   "Carrier_65_Status.3" AT %I3600.3 : Bool;   // POSITIONING_COMPLETE
   "Carrier_65_Status.4" AT %I3600.4 : Bool;   // PRODUCTION HOLD
   "Carrier_65_Status.5" AT %I3600.5 : Bool;   // CARRIER MOVING FORWARD
   "Carrier_65_Status.6" AT %I3600.6 : Bool;   // CARRIER MOVING REVERSE
   "Carrier_65_Status.7" AT %I3600.7 : Bool;   // CARRIER FAULT
   "Carrier_65_Status.8" AT %I3601.0 : Bool;   // CRASH DETECT TRIPPED
   "Carrier_65_Status.9" AT %I3601.1 : Bool;
   "Carrier_65_Status.10" AT %I3601.2 : Bool;
   "Carrier_65_Status.11" AT %I3601.3 : Bool;
   "Carrier_65_Status.12" AT %I3601.4 : Bool;
   "Carrier_65_Status.13" AT %I3601.5 : Bool;
   "Carrier_65_Status.14" AT %I3601.6 : Bool;
   "Carrier_65_Status.15" AT %I3601.7 : Bool;
   "Carrier_65_SDCFaultCode" AT %IW3602 : Word;   // SDC FAULT CODE
   "Carrier_65_CarrierPosition" AT %ID3604 : DWord;   // CARRIER POSITION
   "Carrier_65_CarrierNumber" AT %IW3608 : Word;   // CARRIER NUMBER
   "Carrier_65_G120DControlWord" AT %IW3610 : Word;   // G120D_STW1_CONTROL
   "Carrier_65_G120DControlWord.0" AT %I3610.0 : Bool;   // Bit_00_ON
   "Carrier_65_G120DControlWord.1" AT %I3610.1 : Bool;   // Bit_01_AUS2_INH
   "Carrier_65_G120DControlWord.2" AT %I3610.2 : Bool;   // Bit_02_AUS3_STOP
   "Carrier_65_G120DControlWord.3" AT %I3610.3 : Bool;   // Bit_03_EN
   "Carrier_65_G120DControlWord.4" AT %I3610.4 : Bool;   // Bit_04_EN_RAMP
   "Carrier_65_G120DControlWord.5" AT %I3610.5 : Bool;   // Bit_05_START_RAMP
   "Carrier_65_G120DControlWord.6" AT %I3610.6 : Bool;   // Bit_06_SETPOINT
   "Carrier_65_G120DControlWord.7" AT %I3610.7 : Bool;   // Bit_07_RESET
   "Carrier_65_G120DControlWord.8" AT %I3611.0 : Bool;   // Bit_08_JOG_R
   "Carrier_65_G120DControlWord.9" AT %I3611.1 : Bool;   // Bit_09_JOG_L
   "Carrier_65_G120DControlWord.10" AT %I3611.2 : Bool;   // Bit_10_CONTR_PLC
   "Carrier_65_G120DControlWord.11" AT %I3611.3 : Bool;   // Bit_11_REVERSE
   "Carrier_65_G120DControlWord.12" AT %I3611.4 : Bool;   // Bit_12_BRAKE_RELEASE
   "Carrier_65_G120DControlWord.13" AT %I3611.5 : Bool;   // Bit_13_DDS
   "Carrier_65_G120DControlWord.14" AT %I3611.6 : Bool;   // Bit_14_DO0
   "Carrier_65_G120DControlWord.15" AT %I3611.7 : Bool;   // Bit_15_DO1
   "Carrier_65_G120DStatusWord" AT %IW3612 : Word;   // G120D_ZSW1_STATUS
   "Carrier_65_G120DStatusWord.0" AT %I3612.0 : Bool;   // Bit_00_READY_RUN
   "Carrier_65_G120DStatusWord.1" AT %I3612.1 : Bool;   // Bit_01_READY_ON
   "Carrier_65_G120DStatusWord.2" AT %I3612.2 : Bool;   // Bit_02_ENABLE
   "Carrier_65_G120DStatusWord.3" AT %I3612.3 : Bool;   // Bit_03_FAULT
   "Carrier_65_G120DStatusWord.4" AT %I3612.4 : Bool;   // Bit_04_OFF2
   "Carrier_65_G120DStatusWord.5" AT %I3612.5 : Bool;   // Bit_05_OFF3
   "Carrier_65_G120DStatusWord.6" AT %I3612.6 : Bool;   // Bit_06_LOCK_OUT
   "Carrier_65_G120DStatusWord.7" AT %I3612.7 : Bool;   // Bit_07_WARN
   "Carrier_65_G120DStatusWord.8" AT %I3613.0 : Bool;   // Bit_08_NO_DEVIATION
   "Carrier_65_G120DStatusWord.9" AT %I3613.1 : Bool;   // Bit_09_CONTR_PLC
   "Carrier_65_G120DStatusWord.10" AT %I3613.2 : Bool;   // Bit_10_F_MAX
   "Carrier_65_G120DStatusWord.11" AT %I3613.3 : Bool;   // Bit_11_LIMIT_REACHED
   "Carrier_65_G120DStatusWord.12" AT %I3613.4 : Bool;   // Bit_12_BRAKE_OPEN
   "Carrier_65_G120DStatusWord.13" AT %I3613.5 : Bool;   // Bit_13_NO_OVERTEMP
   "Carrier_65_G120DStatusWord.14" AT %I3613.6 : Bool;   // Bit_14_CW_CCW
   "Carrier_65_G120DStatusWord.15" AT %I3613.7 : Bool;   // Bit_15_OVERL
   "Carrier_65_Slot2_Input" AT %IW3614 : Word;   // SLOT 2 INPUT WORD
   "Carrier_65_CrashDetectSW" AT %I3614.0 : Bool;   // CRASH DETECT SW
   "Carrier_65_SpareSafetyInput(2_1)" AT %I3614.1 : Bool;   // SPARE SAFETY INPUT
   "Carrier_65_SpareSafetyInput(2_2)" AT %I3614.2 : Bool;   // SPARE SAFETY INPUT
   "Carrier_65_SpareSafetyInput(2_3)" AT %I3614.3 : Bool;   // SPARE SAFETY INPUT
   "Carrier_65_SpareSafetyInput(2_4)" AT %I3614.4 : Bool;   // SPARE SAFETY INPUT
   "Carrier_65_SpareSafetyInput(2_5)" AT %I3614.5 : Bool;   // SPARE SAFETY INPUT
   "Carrier_65_SpareSafetyInput(2_6)" AT %I3614.6 : Bool;   // SPARE SAFETY INPUT
   "Carrier_65_SpareSafetyInput(2_7)" AT %I3614.7 : Bool;   // SPARE SAFETY INPUT
   "Carrier_65_Slot3_SafetyOutput" AT %IW3615 : Word;   // SLOT 3 SAFETY OUTPUT WORD
   "Carrier_65_Crash_Detect_OK" AT %I3615.0 : Bool;   // CARRIER CRASH DETECT
   "Carrier_65_SpareSafetyOutput(3_1)" AT %I3615.1 : Bool;   // SPARE SAFETY OUTPUT
   "Carrier_65_SpareSafetyOutput(3_2)" AT %I3615.2 : Bool;   // SPARE SAFETY OUTPUT
   "Carrier_65_SpareSafetyOutput(3_3)" AT %I3615.3 : Bool;   // SPARE SAFETY OUTPUT
   "Carrier_65_SpareSafetyOutput(3_4)" AT %I3615.4 : Bool;   // SPARE SAFETY OUTPUT
   "Carrier_65_SpareSafetyOutput(3_5)" AT %I3615.5 : Bool;   // SPARE SAFETY OUTPUT
   "Carrier_65_SpareSafetyOutput(3_6)" AT %I3615.6 : Bool;   // SPARE SAFETY OUTPUT
   "Carrier_65_SpareSafetyOutput(3_7)" AT %I3615.7 : Bool;   // SPARE SAFETY OUTPUT
   "Carrier_65_Slot4_Input" AT %IW3616 : Word;   // SLOT 4 INPUT WORD
   "Carrier_65_480VPowerOn_MDCB1" AT %I3616.0 : Bool;   // 480 VAC POWER ON MDCB 1
   "Carrier_65_SpareInput(4_1)" AT %I3616.1 : Bool;   // SPARE INPUT
   "Carrier_65_SpareInput(4_2)" AT %I3616.2 : Bool;   // SPARE INPUT
   "Carrier_65_SitopSelectStatus" AT %I3616.3 : Bool;   // SITOP SELECT STATUS
   "Carrier_65_DCsupplyOnPSCB2" AT %I3616.4 : Bool;   // DC SUPPLY ON PSCB 2
   "Carrier_65_SpareInput(4_5)" AT %I3616.5 : Bool;   // SPARE INPUT
   "Carrier_65_SpareInput(4_6)" AT %I3616.6 : Bool;   // SPARE INPUT
   "Carrier_65_SpareInput(4_7)" AT %I3616.7 : Bool;   // SPARE INPUT
   "Carrier_65_PB1_ProdHoldLH" AT %I3617.0 : Bool;   // PB 1 PRODUCTION HOLD LH
   "Carrier_65_PB2_ResetLH" AT %I3617.1 : Bool;   // PB 2 RESET LH
   "Carrier_65_PB3_ProdHoldRH" AT %I3617.2 : Bool;   // PB 3 PRODUCTION HOLD RH
   "Carrier_65_PB4_ResetRH" AT %I3617.3 : Bool;   // PB 4 RESET RH
   "Carrier_65_SpareInput(4_14)" AT %I3617.4 : Bool;   // SPARE INPUT
   "Carrier_65_SpareInput(4_15)" AT %I3617.5 : Bool;   // SPARE INPUT
   "Carrier_65_SpareInput(4_16)" AT %I3617.6 : Bool;   // SPARE INPUT
   "Carrier_65_SpareInput(4_17)" AT %I3617.7 : Bool;   // SPARE INPUT
   "Carrier_65_Slot5_Output" AT %IW3618 : Word;   // SLOT 5 OUTPUT WORD
   "Carrier_65_IRD400_HMI_24VDC_ENABLE" AT %I3618.0 : Bool;   // IRD 400 PANEL HMI 24V DC POWER
   "Carrier_65_FaultLight_LH" AT %I3618.1 : Bool;   // FAULT LIGHT LH
   "Carrier_65_RunLight_LH" AT %I3618.2 : Bool;   // RUN LIGHT LH
   "Carrier_65_FaultLight_RH" AT %I3618.3 : Bool;   // FAULT LIGHT RH
   "Carrier_65_RunLight_RH" AT %I3618.4 : Bool;   // RUN LIGHT RH
   "Carrier_65_SpareOutput(5_5)" AT %I3618.5 : Bool;   // SPARE OUTPUT
   "Carrier_65_SpareOutput(5_6)" AT %I3618.6 : Bool;   // SPARE OUTPUT
   "Carrier_65_SpareOutput(5_7)" AT %I3618.7 : Bool;   // SPARE OUTPUT
   "Carrier_65_ActualSpeed" AT %IW3620 : Word;   // ACTUAL SPEED
   "Carrier_65_CarrierDriveAlarm" AT %IW3622 : Word;   // CARRIER DRIVE ALARM
   "Carrier_65_CarrierDriveWarning" AT %IW3624 : Word;   // CARRIER DRIVE WARNING
   "Carrier_66_Status" AT %IW3650 : Word;   // CARRIER STATUS WORD
   "Carrier_66_Status.0" AT %I3650.0 : Bool;   // HEARTBEAT
   "Carrier_66_Status.1" AT %I3650.1 : Bool;   // MANUAL
   "Carrier_66_Status.2" AT %I3650.2 : Bool;   // IN_AUTO
   "Carrier_66_Status.3" AT %I3650.3 : Bool;   // POSITIONING_COMPLETE
   "Carrier_66_Status.4" AT %I3650.4 : Bool;   // PRODUCTION HOLD
   "Carrier_66_Status.5" AT %I3650.5 : Bool;   // CARRIER MOVING FORWARD
   "Carrier_66_Status.6" AT %I3650.6 : Bool;   // CARRIER MOVING REVERSE
   "Carrier_66_Status.7" AT %I3650.7 : Bool;   // CARRIER FAULT
   "Carrier_66_Status.8" AT %I3651.0 : Bool;   // CRASH DETECT TRIPPED
   "Carrier_66_Status.9" AT %I3651.1 : Bool;
   "Carrier_66_Status.10" AT %I3651.2 : Bool;
   "Carrier_66_Status.11" AT %I3651.3 : Bool;
   "Carrier_66_Status.12" AT %I3651.4 : Bool;
   "Carrier_66_Status.13" AT %I3651.5 : Bool;
   "Carrier_66_Status.14" AT %I3651.6 : Bool;
   "Carrier_66_Status.15" AT %I3651.7 : Bool;
   "Carrier_66_SDCFaultCode" AT %IW3652 : Word;   // SDC FAULT CODE
   "Carrier_66_CarrierPosition" AT %ID3654 : DWord;   // CARRIER POSITION
   "Carrier_66_CarrierNumber" AT %IW3658 : Word;   // CARRIER NUMBER
   "Carrier_66_G120DControlWord" AT %IW3660 : Word;   // G120D_STW1_CONTROL
   "Carrier_66_G120DControlWord.0" AT %I3660.0 : Bool;   // Bit_00_ON
   "Carrier_66_G120DControlWord.1" AT %I3660.1 : Bool;   // Bit_01_AUS2_INH
   "Carrier_66_G120DControlWord.2" AT %I3660.2 : Bool;   // Bit_02_AUS3_STOP
   "Carrier_66_G120DControlWord.3" AT %I3660.3 : Bool;   // Bit_03_EN
   "Carrier_66_G120DControlWord.4" AT %I3660.4 : Bool;   // Bit_04_EN_RAMP
   "Carrier_66_G120DControlWord.5" AT %I3660.5 : Bool;   // Bit_05_START_RAMP
   "Carrier_66_G120DControlWord.6" AT %I3660.6 : Bool;   // Bit_06_SETPOINT
   "Carrier_66_G120DControlWord.7" AT %I3660.7 : Bool;   // Bit_07_RESET
   "Carrier_66_G120DControlWord.8" AT %I3661.0 : Bool;   // Bit_08_JOG_R
   "Carrier_66_G120DControlWord.9" AT %I3661.1 : Bool;   // Bit_09_JOG_L
   "Carrier_66_G120DControlWord.10" AT %I3661.2 : Bool;   // Bit_10_CONTR_PLC
   "Carrier_66_G120DControlWord.11" AT %I3661.3 : Bool;   // Bit_11_REVERSE
   "Carrier_66_G120DControlWord.12" AT %I3661.4 : Bool;   // Bit_12_BRAKE_RELEASE
   "Carrier_66_G120DControlWord.13" AT %I3661.5 : Bool;   // Bit_13_DDS
   "Carrier_66_G120DControlWord.14" AT %I3661.6 : Bool;   // Bit_14_DO0
   "Carrier_66_G120DControlWord.15" AT %I3661.7 : Bool;   // Bit_15_DO1
   "Carrier_66_G120DStatusWord" AT %IW3662 : Word;   // G120D_ZSW1_STATUS
   "Carrier_66_G120DStatusWord.0" AT %I3662.0 : Bool;   // Bit_00_READY_RUN
   "Carrier_66_G120DStatusWord.1" AT %I3662.1 : Bool;   // Bit_01_READY_ON
   "Carrier_66_G120DStatusWord.2" AT %I3662.2 : Bool;   // Bit_02_ENABLE
   "Carrier_66_G120DStatusWord.3" AT %I3662.3 : Bool;   // Bit_03_FAULT
   "Carrier_66_G120DStatusWord.4" AT %I3662.4 : Bool;   // Bit_04_OFF2
   "Carrier_66_G120DStatusWord.5" AT %I3662.5 : Bool;   // Bit_05_OFF3
   "Carrier_66_G120DStatusWord.6" AT %I3662.6 : Bool;   // Bit_06_LOCK_OUT
   "Carrier_66_G120DStatusWord.7" AT %I3662.7 : Bool;   // Bit_07_WARN
   "Carrier_66_G120DStatusWord.8" AT %I3663.0 : Bool;   // Bit_08_NO_DEVIATION
   "Carrier_66_G120DStatusWord.9" AT %I3663.1 : Bool;   // Bit_09_CONTR_PLC
   "Carrier_66_G120DStatusWord.10" AT %I3663.2 : Bool;   // Bit_10_F_MAX
   "Carrier_66_G120DStatusWord.11" AT %I3663.3 : Bool;   // Bit_11_LIMIT_REACHED
   "Carrier_66_G120DStatusWord.12" AT %I3663.4 : Bool;   // Bit_12_BRAKE_OPEN
   "Carrier_66_G120DStatusWord.13" AT %I3663.5 : Bool;   // Bit_13_NO_OVERTEMP
   "Carrier_66_G120DStatusWord.14" AT %I3663.6 : Bool;   // Bit_14_CW_CCW
   "Carrier_66_G120DStatusWord.15" AT %I3663.7 : Bool;   // Bit_15_OVERL
   "Carrier_66_Slot2_Input" AT %IW3664 : Word;   // SLOT 2 INPUT WORD
   "Carrier_66_CrashDetectSW" AT %I3664.0 : Bool;   // CRASH DETECT SW
   "Carrier_66_SpareSafetyInput(2_1)" AT %I3664.1 : Bool;   // SPARE SAFETY INPUT
   "Carrier_66_SpareSafetyInput(2_2)" AT %I3664.2 : Bool;   // SPARE SAFETY INPUT
   "Carrier_66_SpareSafetyInput(2_3)" AT %I3664.3 : Bool;   // SPARE SAFETY INPUT
   "Carrier_66_SpareSafetyInput(2_4)" AT %I3664.4 : Bool;   // SPARE SAFETY INPUT
   "Carrier_66_SpareSafetyInput(2_5)" AT %I3664.5 : Bool;   // SPARE SAFETY INPUT
   "Carrier_66_SpareSafetyInput(2_6)" AT %I3664.6 : Bool;   // SPARE SAFETY INPUT
   "Carrier_66_SpareSafetyInput(2_7)" AT %I3664.7 : Bool;   // SPARE SAFETY INPUT
   "Carrier_66_Slot3_SafetyOutput" AT %IW3665 : Word;   // SLOT 3 SAFETY OUTPUT WORD
   "Carrier_66_Crash_Detect_OK" AT %I3665.0 : Bool;   // CARRIER CRASH DETECT
   "Carrier_66_SpareSafetyOutput(3_1)" AT %I3665.1 : Bool;   // SPARE SAFETY OUTPUT
   "Carrier_66_SpareSafetyOutput(3_2)" AT %I3665.2 : Bool;   // SPARE SAFETY OUTPUT
   "Carrier_66_SpareSafetyOutput(3_3)" AT %I3665.3 : Bool;   // SPARE SAFETY OUTPUT
   "Carrier_66_SpareSafetyOutput(3_4)" AT %I3665.4 : Bool;   // SPARE SAFETY OUTPUT
   "Carrier_66_SpareSafetyOutput(3_5)" AT %I3665.5 : Bool;   // SPARE SAFETY OUTPUT
   "Carrier_66_SpareSafetyOutput(3_6)" AT %I3665.6 : Bool;   // SPARE SAFETY OUTPUT
   "Carrier_66_SpareSafetyOutput(3_7)" AT %I3665.7 : Bool;   // SPARE SAFETY OUTPUT
   "Carrier_66_Slot4_Input" AT %IW3666 : Word;   // SLOT 4 INPUT WORD
   "Carrier_66_480VPowerOn_MDCB1" AT %I3666.0 : Bool;   // 480 VAC POWER ON MDCB 1
   "Carrier_66_SpareInput(4_1)" AT %I3666.1 : Bool;   // SPARE INPUT
   "Carrier_66_SpareInput(4_2)" AT %I3666.2 : Bool;   // SPARE INPUT
   "Carrier_66_SitopSelectStatus" AT %I3666.3 : Bool;   // SITOP SELECT STATUS
   "Carrier_66_DCsupplyOnPSCB2" AT %I3666.4 : Bool;   // DC SUPPLY ON PSCB 2
   "Carrier_66_SpareInput(4_5)" AT %I3666.5 : Bool;   // SPARE INPUT
   "Carrier_66_SpareInput(4_6)" AT %I3666.6 : Bool;   // SPARE INPUT
   "Carrier_66_SpareInput(4_7)" AT %I3666.7 : Bool;   // SPARE INPUT
   "Carrier_66_PB1_ProdHoldLH" AT %I3667.0 : Bool;   // PB 1 PRODUCTION HOLD LH
   "Carrier_66_PB2_ResetLH" AT %I3667.1 : Bool;   // PB 2 RESET LH
   "Carrier_66_PB3_ProdHoldRH" AT %I3667.2 : Bool;   // PB 3 PRODUCTION HOLD RH
   "Carrier_66_PB4_ResetRH" AT %I3667.3 : Bool;   // PB 4 RESET RH
   "Carrier_66_SpareInput(4_14)" AT %I3667.4 : Bool;   // SPARE INPUT
   "Carrier_66_SpareInput(4_15)" AT %I3667.5 : Bool;   // SPARE INPUT
   "Carrier_66_SpareInput(4_16)" AT %I3667.6 : Bool;   // SPARE INPUT
   "Carrier_66_SpareInput(4_17)" AT %I3667.7 : Bool;   // SPARE INPUT
   "Carrier_66_Slot5_Output" AT %IW3668 : Word;   // SLOT 5 OUTPUT WORD
   "Carrier_66_IRD400_HMI_24VDC_ENABLE" AT %I3668.0 : Bool;   // IRD 400 PANEL HMI 24V DC POWER
   "Carrier_66_FaultLight_LH" AT %I3668.1 : Bool;   // FAULT LIGHT LH
   "Carrier_66_RunLight_LH" AT %I3668.2 : Bool;   // RUN LIGHT LH
   "Carrier_66_FaultLight_RH" AT %I3668.3 : Bool;   // FAULT LIGHT RH
   "Carrier_66_RunLight_RH" AT %I3668.4 : Bool;   // RUN LIGHT RH
   "Carrier_66_SpareOutput(5_5)" AT %I3668.5 : Bool;   // SPARE OUTPUT
   "Carrier_66_SpareOutput(5_6)" AT %I3668.6 : Bool;   // SPARE OUTPUT
   "Carrier_66_SpareOutput(5_7)" AT %I3668.7 : Bool;   // SPARE OUTPUT
   "Carrier_66_ActualSpeed" AT %IW3670 : Word;   // ACTUAL SPEED
   "Carrier_66_CarrierDriveAlarm" AT %IW3672 : Word;   // CARRIER DRIVE ALARM
   "Carrier_66_CarrierDriveWarning" AT %IW3674 : Word;   // CARRIER DRIVE WARNING
   "Carrier_67_Status" AT %IW3700 : Word;   // CARRIER STATUS WORD
   "Carrier_67_Status.0" AT %I3700.0 : Bool;   // HEARTBEAT
   "Carrier_67_Status.1" AT %I3700.1 : Bool;   // MANUAL
   "Carrier_67_Status.2" AT %I3700.2 : Bool;   // IN_AUTO
   "Carrier_67_Status.3" AT %I3700.3 : Bool;   // POSITIONING_COMPLETE
   "Carrier_67_Status.4" AT %I3700.4 : Bool;   // PRODUCTION HOLD
   "Carrier_67_Status.5" AT %I3700.5 : Bool;   // CARRIER MOVING FORWARD
   "Carrier_67_Status.6" AT %I3700.6 : Bool;   // CARRIER MOVING REVERSE
   "Carrier_67_Status.7" AT %I3700.7 : Bool;   // CARRIER FAULT
   "Carrier_67_Status.8" AT %I3701.0 : Bool;   // CRASH DETECT TRIPPED
   "Carrier_67_Status.9" AT %I3701.1 : Bool;
   "Carrier_67_Status.10" AT %I3701.2 : Bool;
   "Carrier_67_Status.11" AT %I3701.3 : Bool;
   "Carrier_67_Status.12" AT %I3701.4 : Bool;
   "Carrier_67_Status.13" AT %I3701.5 : Bool;
   "Carrier_67_Status.14" AT %I3701.6 : Bool;
   "Carrier_67_Status.15" AT %I3701.7 : Bool;
   "Carrier_67_SDCFaultCode" AT %IW3702 : Word;   // SDC FAULT CODE
   "Carrier_67_CarrierPosition" AT %ID3704 : DWord;   // CARRIER POSITION
   "Carrier_67_CarrierNumber" AT %IW3708 : Word;   // CARRIER NUMBER
   "Carrier_67_G120DControlWord" AT %IW3710 : Word;   // G120D_STW1_CONTROL
   "Carrier_67_G120DControlWord.0" AT %I3710.0 : Bool;   // Bit_00_ON
   "Carrier_67_G120DControlWord.1" AT %I3710.1 : Bool;   // Bit_01_AUS2_INH
   "Carrier_67_G120DControlWord.2" AT %I3710.2 : Bool;   // Bit_02_AUS3_STOP
   "Carrier_67_G120DControlWord.3" AT %I3710.3 : Bool;   // Bit_03_EN
   "Carrier_67_G120DControlWord.4" AT %I3710.4 : Bool;   // Bit_04_EN_RAMP
   "Carrier_67_G120DControlWord.5" AT %I3710.5 : Bool;   // Bit_05_START_RAMP
   "Carrier_67_G120DControlWord.6" AT %I3710.6 : Bool;   // Bit_06_SETPOINT
   "Carrier_67_G120DControlWord.7" AT %I3710.7 : Bool;   // Bit_07_RESET
   "Carrier_67_G120DControlWord.8" AT %I3711.0 : Bool;   // Bit_08_JOG_R
   "Carrier_67_G120DControlWord.9" AT %I3711.1 : Bool;   // Bit_09_JOG_L
   "Carrier_67_G120DControlWord.10" AT %I3711.2 : Bool;   // Bit_10_CONTR_PLC
   "Carrier_67_G120DControlWord.11" AT %I3711.3 : Bool;   // Bit_11_REVERSE
   "Carrier_67_G120DControlWord.12" AT %I3711.4 : Bool;   // Bit_12_BRAKE_RELEASE
   "Carrier_67_G120DControlWord.13" AT %I3711.5 : Bool;   // Bit_13_DDS
   "Carrier_67_G120DControlWord.14" AT %I3711.6 : Bool;   // Bit_14_DO0
   "Carrier_67_G120DControlWord.15" AT %I3711.7 : Bool;   // Bit_15_DO1
   "Carrier_67_G120DStatusWord" AT %IW3712 : Word;   // G120D_ZSW1_STATUS
   "Carrier_67_G120DStatusWord.0" AT %I3712.0 : Bool;   // Bit_00_READY_RUN
   "Carrier_67_G120DStatusWord.1" AT %I3712.1 : Bool;   // Bit_01_READY_ON
   "Carrier_67_G120DStatusWord.2" AT %I3712.2 : Bool;   // Bit_02_ENABLE
   "Carrier_67_G120DStatusWord.3" AT %I3712.3 : Bool;   // Bit_03_FAULT
   "Carrier_67_G120DStatusWord.4" AT %I3712.4 : Bool;   // Bit_04_OFF2
   "Carrier_67_G120DStatusWord.5" AT %I3712.5 : Bool;   // Bit_05_OFF3
   "Carrier_67_G120DStatusWord.6" AT %I3712.6 : Bool;   // Bit_06_LOCK_OUT
   "Carrier_67_G120DStatusWord.7" AT %I3712.7 : Bool;   // Bit_07_WARN
   "Carrier_67_G120DStatusWord.8" AT %I3713.0 : Bool;   // Bit_08_NO_DEVIATION
   "Carrier_67_G120DStatusWord.9" AT %I3713.1 : Bool;   // Bit_09_CONTR_PLC
   "Carrier_67_G120DStatusWord.10" AT %I3713.2 : Bool;   // Bit_10_F_MAX
   "Carrier_67_G120DStatusWord.11" AT %I3713.3 : Bool;   // Bit_11_LIMIT_REACHED
   "Carrier_67_G120DStatusWord.12" AT %I3713.4 : Bool;   // Bit_12_BRAKE_OPEN
   "Carrier_67_G120DStatusWord.13" AT %I3713.5 : Bool;   // Bit_13_NO_OVERTEMP
   "Carrier_67_G120DStatusWord.14" AT %I3713.6 : Bool;   // Bit_14_CW_CCW
   "Carrier_67_G120DStatusWord.15" AT %I3713.7 : Bool;   // Bit_15_OVERL
   "Carrier_67_Slot2_Input" AT %IW3714 : Word;   // SLOT 2 INPUT WORD
   "Carrier_67_CrashDetectSW" AT %I3714.0 : Bool;   // CRASH DETECT SW
   "Carrier_67_SpareSafetyInput(2_1)" AT %I3714.1 : Bool;   // SPARE SAFETY INPUT
   "Carrier_67_SpareSafetyInput(2_2)" AT %I3714.2 : Bool;   // SPARE SAFETY INPUT
   "Carrier_67_SpareSafetyInput(2_3)" AT %I3714.3 : Bool;   // SPARE SAFETY INPUT
   "Carrier_67_SpareSafetyInput(2_4)" AT %I3714.4 : Bool;   // SPARE SAFETY INPUT
   "Carrier_67_SpareSafetyInput(2_5)" AT %I3714.5 : Bool;   // SPARE SAFETY INPUT
   "Carrier_67_SpareSafetyInput(2_6)" AT %I3714.6 : Bool;   // SPARE SAFETY INPUT
   "Carrier_67_SpareSafetyInput(2_7)" AT %I3714.7 : Bool;   // SPARE SAFETY INPUT
   "Carrier_67_Slot3_SafetyOutput" AT %IW3715 : Word;   // SLOT 3 SAFETY OUTPUT WORD
   "Carrier_67_Crash_Detect_OK" AT %I3715.0 : Bool;   // CARRIER CRASH DETECT
   "Carrier_67_SpareSafetyOutput(3_1)" AT %I3715.1 : Bool;   // SPARE SAFETY OUTPUT
   "Carrier_67_SpareSafetyOutput(3_2)" AT %I3715.2 : Bool;   // SPARE SAFETY OUTPUT
   "Carrier_67_SpareSafetyOutput(3_3)" AT %I3715.3 : Bool;   // SPARE SAFETY OUTPUT
   "Carrier_67_SpareSafetyOutput(3_4)" AT %I3715.4 : Bool;   // SPARE SAFETY OUTPUT
   "Carrier_67_SpareSafetyOutput(3_5)" AT %I3715.5 : Bool;   // SPARE SAFETY OUTPUT
   "Carrier_67_SpareSafetyOutput(3_6)" AT %I3715.6 : Bool;   // SPARE SAFETY OUTPUT
   "Carrier_67_SpareSafetyOutput(3_7)" AT %I3715.7 : Bool;   // SPARE SAFETY OUTPUT
   "Carrier_67_Slot4_Input" AT %IW3716 : Word;   // SLOT 4 INPUT WORD
   "Carrier_67_480VPowerOn_MDCB1" AT %I3716.0 : Bool;   // 480 VAC POWER ON MDCB 1
   "Carrier_67_SpareInput(4_1)" AT %I3716.1 : Bool;   // SPARE INPUT
   "Carrier_67_SpareInput(4_2)" AT %I3716.2 : Bool;   // SPARE INPUT
   "Carrier_67_SitopSelectStatus" AT %I3716.3 : Bool;   // SITOP SELECT STATUS
   "Carrier_67_DCsupplyOnPSCB2" AT %I3716.4 : Bool;   // DC SUPPLY ON PSCB 2
   "Carrier_67_SpareInput(4_5)" AT %I3716.5 : Bool;   // SPARE INPUT
   "Carrier_67_SpareInput(4_6)" AT %I3716.6 : Bool;   // SPARE INPUT
   "Carrier_67_SpareInput(4_7)" AT %I3716.7 : Bool;   // SPARE INPUT
   "Carrier_67_PB1_ProdHoldLH" AT %I3717.0 : Bool;   // PB 1 PRODUCTION HOLD LH
   "Carrier_67_PB2_ResetLH" AT %I3717.1 : Bool;   // PB 2 RESET LH
   "Carrier_67_PB3_ProdHoldRH" AT %I3717.2 : Bool;   // PB 3 PRODUCTION HOLD RH
   "Carrier_67_PB4_ResetRH" AT %I3717.3 : Bool;   // PB 4 RESET RH
   "Carrier_67_SpareInput(4_14)" AT %I3717.4 : Bool;   // SPARE INPUT
   "Carrier_67_SpareInput(4_15)" AT %I3717.5 : Bool;   // SPARE INPUT
   "Carrier_67_SpareInput(4_16)" AT %I3717.6 : Bool;   // SPARE INPUT
   "Carrier_67_SpareInput(4_17)" AT %I3717.7 : Bool;   // SPARE INPUT
   "Carrier_67_Slot5_Output" AT %IW3718 : Word;   // SLOT 5 OUTPUT WORD
   "Carrier_67_IRD400_HMI_24VDC_ENABLE" AT %I3718.0 : Bool;   // IRD 400 PANEL HMI 24V DC POWER
   "Carrier_67_FaultLight_LH" AT %I3718.1 : Bool;   // FAULT LIGHT LH
   "Carrier_67_RunLight_LH" AT %I3718.2 : Bool;   // RUN LIGHT LH
   "Carrier_67_FaultLight_RH" AT %I3718.3 : Bool;   // FAULT LIGHT RH
   "Carrier_67_RunLight_RH" AT %I3718.4 : Bool;   // RUN LIGHT RH
   "Carrier_67_SpareOutput(5_5)" AT %I3718.5 : Bool;   // SPARE OUTPUT
   "Carrier_67_SpareOutput(5_6)" AT %I3718.6 : Bool;   // SPARE OUTPUT
   "Carrier_67_SpareOutput(5_7)" AT %I3718.7 : Bool;   // SPARE OUTPUT
   "Carrier_67_ActualSpeed" AT %IW3720 : Word;   // ACTUAL SPEED
   "Carrier_67_CarrierDriveAlarm" AT %IW3722 : Word;   // CARRIER DRIVE ALARM
   "Carrier_67_CarrierDriveWarning" AT %IW3724 : Word;   // CARRIER DRIVE WARNING
   "Carrier_68_Status" AT %IW3750 : Word;   // CARRIER STATUS WORD
   "Carrier_68_Status.0" AT %I3750.0 : Bool;   // HEARTBEAT
   "Carrier_68_Status.1" AT %I3750.1 : Bool;   // MANUAL
   "Carrier_68_Status.2" AT %I3750.2 : Bool;   // IN_AUTO
   "Carrier_68_Status.3" AT %I3750.3 : Bool;   // POSITIONING_COMPLETE
   "Carrier_68_Status.4" AT %I3750.4 : Bool;   // PRODUCTION HOLD
   "Carrier_68_Status.5" AT %I3750.5 : Bool;   // CARRIER MOVING FORWARD
   "Carrier_68_Status.6" AT %I3750.6 : Bool;   // CARRIER MOVING REVERSE
   "Carrier_68_Status.7" AT %I3750.7 : Bool;   // CARRIER FAULT
   "Carrier_68_Status.8" AT %I3751.0 : Bool;   // CRASH DETECT TRIPPED
   "Carrier_68_Status.9" AT %I3751.1 : Bool;
   "Carrier_68_Status.10" AT %I3751.2 : Bool;
   "Carrier_68_Status.11" AT %I3751.3 : Bool;
   "Carrier_68_Status.12" AT %I3751.4 : Bool;
   "Carrier_68_Status.13" AT %I3751.5 : Bool;
   "Carrier_68_Status.14" AT %I3751.6 : Bool;
   "Carrier_68_Status.15" AT %I3751.7 : Bool;
   "Carrier_68_SDCFaultCode" AT %IW3752 : Word;   // SDC FAULT CODE
   "Carrier_68_CarrierPosition" AT %ID3754 : DWord;   // CARRIER POSITION
   "Carrier_68_CarrierNumber" AT %IW3758 : Word;   // CARRIER NUMBER
   "Carrier_68_G120DControlWord" AT %IW3760 : Word;   // G120D_STW1_CONTROL
   "Carrier_68_G120DControlWord.0" AT %I3760.0 : Bool;   // Bit_00_ON
   "Carrier_68_G120DControlWord.1" AT %I3760.1 : Bool;   // Bit_01_AUS2_INH
   "Carrier_68_G120DControlWord.2" AT %I3760.2 : Bool;   // Bit_02_AUS3_STOP
   "Carrier_68_G120DControlWord.3" AT %I3760.3 : Bool;   // Bit_03_EN
   "Carrier_68_G120DControlWord.4" AT %I3760.4 : Bool;   // Bit_04_EN_RAMP
   "Carrier_68_G120DControlWord.5" AT %I3760.5 : Bool;   // Bit_05_START_RAMP
   "Carrier_68_G120DControlWord.6" AT %I3760.6 : Bool;   // Bit_06_SETPOINT
   "Carrier_68_G120DControlWord.7" AT %I3760.7 : Bool;   // Bit_07_RESET
   "Carrier_68_G120DControlWord.8" AT %I3761.0 : Bool;   // Bit_08_JOG_R
   "Carrier_68_G120DControlWord.9" AT %I3761.1 : Bool;   // Bit_09_JOG_L
   "Carrier_68_G120DControlWord.10" AT %I3761.2 : Bool;   // Bit_10_CONTR_PLC
   "Carrier_68_G120DControlWord.11" AT %I3761.3 : Bool;   // Bit_11_REVERSE
   "Carrier_68_G120DControlWord.12" AT %I3761.4 : Bool;   // Bit_12_BRAKE_RELEASE
   "Carrier_68_G120DControlWord.13" AT %I3761.5 : Bool;   // Bit_13_DDS
   "Carrier_68_G120DControlWord.14" AT %I3761.6 : Bool;   // Bit_14_DO0
   "Carrier_68_G120DControlWord.15" AT %I3761.7 : Bool;   // Bit_15_DO1
   "Carrier_68_G120DStatusWord" AT %IW3762 : Word;   // G120D_ZSW1_STATUS
   "Carrier_68_G120DStatusWord.0" AT %I3762.0 : Bool;   // Bit_00_READY_RUN
   "Carrier_68_G120DStatusWord.1" AT %I3762.1 : Bool;   // Bit_01_READY_ON
   "Carrier_68_G120DStatusWord.2" AT %I3762.2 : Bool;   // Bit_02_ENABLE
   "Carrier_68_G120DStatusWord.3" AT %I3762.3 : Bool;   // Bit_03_FAULT
   "Carrier_68_G120DStatusWord.4" AT %I3762.4 : Bool;   // Bit_04_OFF2
   "Carrier_68_G120DStatusWord.5" AT %I3762.5 : Bool;   // Bit_05_OFF3
   "Carrier_68_G120DStatusWord.6" AT %I3762.6 : Bool;   // Bit_06_LOCK_OUT
   "Carrier_68_G120DStatusWord.7" AT %I3762.7 : Bool;   // Bit_07_WARN
   "Carrier_68_G120DStatusWord.8" AT %I3763.0 : Bool;   // Bit_08_NO_DEVIATION
   "Carrier_68_G120DStatusWord.9" AT %I3763.1 : Bool;   // Bit_09_CONTR_PLC
   "Carrier_68_G120DStatusWord.10" AT %I3763.2 : Bool;   // Bit_10_F_MAX
   "Carrier_68_G120DStatusWord.11" AT %I3763.3 : Bool;   // Bit_11_LIMIT_REACHED
   "Carrier_68_G120DStatusWord.12" AT %I3763.4 : Bool;   // Bit_12_BRAKE_OPEN
   "Carrier_68_G120DStatusWord.13" AT %I3763.5 : Bool;   // Bit_13_NO_OVERTEMP
   "Carrier_68_G120DStatusWord.14" AT %I3763.6 : Bool;   // Bit_14_CW_CCW
   "Carrier_68_G120DStatusWord.15" AT %I3763.7 : Bool;   // Bit_15_OVERL
   "Carrier_68_Slot2_Input" AT %IW3764 : Word;   // SLOT 2 INPUT WORD
   "Carrier_68_CrashDetectSW" AT %I3764.0 : Bool;   // CRASH DETECT SW
   "Carrier_68_SpareSafetyInput(2_1)" AT %I3764.1 : Bool;   // SPARE SAFETY INPUT
   "Carrier_68_SpareSafetyInput(2_2)" AT %I3764.2 : Bool;   // SPARE SAFETY INPUT
   "Carrier_68_SpareSafetyInput(2_3)" AT %I3764.3 : Bool;   // SPARE SAFETY INPUT
   "Carrier_68_SpareSafetyInput(2_4)" AT %I3764.4 : Bool;   // SPARE SAFETY INPUT
   "Carrier_68_SpareSafetyInput(2_5)" AT %I3764.5 : Bool;   // SPARE SAFETY INPUT
   "Carrier_68_SpareSafetyInput(2_6)" AT %I3764.6 : Bool;   // SPARE SAFETY INPUT
   "Carrier_68_SpareSafetyInput(2_7)" AT %I3764.7 : Bool;   // SPARE SAFETY INPUT
   "Carrier_68_Slot3_SafetyOutput" AT %IW3765 : Word;   // SLOT 3 SAFETY OUTPUT WORD
   "Carrier_68_Crash_Detect_OK" AT %I3765.0 : Bool;   // CARRIER CRASH DETECT
   "Carrier_68_SpareSafetyOutput(3_1)" AT %I3765.1 : Bool;   // SPARE SAFETY OUTPUT
   "Carrier_68_SpareSafetyOutput(3_2)" AT %I3765.2 : Bool;   // SPARE SAFETY OUTPUT
   "Carrier_68_SpareSafetyOutput(3_3)" AT %I3765.3 : Bool;   // SPARE SAFETY OUTPUT
   "Carrier_68_SpareSafetyOutput(3_4)" AT %I3765.4 : Bool;   // SPARE SAFETY OUTPUT
   "Carrier_68_SpareSafetyOutput(3_5)" AT %I3765.5 : Bool;   // SPARE SAFETY OUTPUT
   "Carrier_68_SpareSafetyOutput(3_6)" AT %I3765.6 : Bool;   // SPARE SAFETY OUTPUT
   "Carrier_68_SpareSafetyOutput(3_7)" AT %I3765.7 : Bool;   // SPARE SAFETY OUTPUT
   "Carrier_68_Slot4_Input" AT %IW3766 : Word;   // SLOT 4 INPUT WORD
   "Carrier_68_480VPowerOn_MDCB1" AT %I3766.0 : Bool;   // 480 VAC POWER ON MDCB 1
   "Carrier_68_SpareInput(4_1)" AT %I3766.1 : Bool;   // SPARE INPUT
   "Carrier_68_SpareInput(4_2)" AT %I3766.2 : Bool;   // SPARE INPUT
   "Carrier_68_SitopSelectStatus" AT %I3766.3 : Bool;   // SITOP SELECT STATUS
   "Carrier_68_DCsupplyOnPSCB2" AT %I3766.4 : Bool;   // DC SUPPLY ON PSCB 2
   "Carrier_68_SpareInput(4_5)" AT %I3766.5 : Bool;   // SPARE INPUT
   "Carrier_68_SpareInput(4_6)" AT %I3766.6 : Bool;   // SPARE INPUT
   "Carrier_68_SpareInput(4_7)" AT %I3766.7 : Bool;   // SPARE INPUT
   "Carrier_68_PB1_ProdHoldLH" AT %I3767.0 : Bool;   // PB 1 PRODUCTION HOLD LH
   "Carrier_68_PB2_ResetLH" AT %I3767.1 : Bool;   // PB 2 RESET LH
   "Carrier_68_PB3_ProdHoldRH" AT %I3767.2 : Bool;   // PB 3 PRODUCTION HOLD RH
   "Carrier_68_PB4_ResetRH" AT %I3767.3 : Bool;   // PB 4 RESET RH
   "Carrier_68_SpareInput(4_14)" AT %I3767.4 : Bool;   // SPARE INPUT
   "Carrier_68_SpareInput(4_15)" AT %I3767.5 : Bool;   // SPARE INPUT
   "Carrier_68_SpareInput(4_16)" AT %I3767.6 : Bool;   // SPARE INPUT
   "Carrier_68_SpareInput(4_17)" AT %I3767.7 : Bool;   // SPARE INPUT
   "Carrier_68_Slot5_Output" AT %IW3768 : Word;   // SLOT 5 OUTPUT WORD
   "Carrier_68_IRD400_HMI_24VDC_ENABLE" AT %I3768.0 : Bool;   // IRD 400 PANEL HMI 24V DC POWER
   "Carrier_68_FaultLight_LH" AT %I3768.1 : Bool;   // FAULT LIGHT LH
   "Carrier_68_RunLight_LH" AT %I3768.2 : Bool;   // RUN LIGHT LH
   "Carrier_68_FaultLight_RH" AT %I3768.3 : Bool;   // FAULT LIGHT RH
   "Carrier_68_RunLight_RH" AT %I3768.4 : Bool;   // RUN LIGHT RH
   "Carrier_68_SpareOutput(5_5)" AT %I3768.5 : Bool;   // SPARE OUTPUT
   "Carrier_68_SpareOutput(5_6)" AT %I3768.6 : Bool;   // SPARE OUTPUT
   "Carrier_68_SpareOutput(5_7)" AT %I3768.7 : Bool;   // SPARE OUTPUT
   "Carrier_68_ActualSpeed" AT %IW3770 : Word;   // ACTUAL SPEED
   "Carrier_68_CarrierDriveAlarm" AT %IW3772 : Word;   // CARRIER DRIVE ALARM
   "Carrier_68_CarrierDriveWarning" AT %IW3774 : Word;   // CARRIER DRIVE WARNING
   "Carrier_69_Status" AT %IW3800 : Word;   // CARRIER STATUS WORD
   "Carrier_69_Status.0" AT %I3800.0 : Bool;   // HEARTBEAT
   "Carrier_69_Status.1" AT %I3800.1 : Bool;   // MANUAL
   "Carrier_69_Status.2" AT %I3800.2 : Bool;   // IN_AUTO
   "Carrier_69_Status.3" AT %I3800.3 : Bool;   // POSITIONING_COMPLETE
   "Carrier_69_Status.4" AT %I3800.4 : Bool;   // PRODUCTION HOLD
   "Carrier_69_Status.5" AT %I3800.5 : Bool;   // CARRIER MOVING FORWARD
   "Carrier_69_Status.6" AT %I3800.6 : Bool;   // CARRIER MOVING REVERSE
   "Carrier_69_Status.7" AT %I3800.7 : Bool;   // CARRIER FAULT
   "Carrier_69_Status.8" AT %I3801.0 : Bool;   // CRASH DETECT TRIPPED
   "Carrier_69_Status.9" AT %I3801.1 : Bool;
   "Carrier_69_Status.10" AT %I3801.2 : Bool;
   "Carrier_69_Status.11" AT %I3801.3 : Bool;
   "Carrier_69_Status.12" AT %I3801.4 : Bool;
   "Carrier_69_Status.13" AT %I3801.5 : Bool;
   "Carrier_69_Status.14" AT %I3801.6 : Bool;
   "Carrier_69_Status.15" AT %I3801.7 : Bool;
   "Carrier_69_SDCFaultCode" AT %IW3802 : Word;   // SDC FAULT CODE
   "Carrier_69_CarrierPosition" AT %ID3804 : DWord;   // CARRIER POSITION
   "Carrier_69_CarrierNumber" AT %IW3808 : Word;   // CARRIER NUMBER
   "Carrier_69_G120DControlWord" AT %IW3810 : Word;   // G120D_STW1_CONTROL
   "Carrier_69_G120DControlWord.0" AT %I3810.0 : Bool;   // Bit_00_ON
   "Carrier_69_G120DControlWord.1" AT %I3810.1 : Bool;   // Bit_01_AUS2_INH
   "Carrier_69_G120DControlWord.2" AT %I3810.2 : Bool;   // Bit_02_AUS3_STOP
   "Carrier_69_G120DControlWord.3" AT %I3810.3 : Bool;   // Bit_03_EN
   "Carrier_69_G120DControlWord.4" AT %I3810.4 : Bool;   // Bit_04_EN_RAMP
   "Carrier_69_G120DControlWord.5" AT %I3810.5 : Bool;   // Bit_05_START_RAMP
   "Carrier_69_G120DControlWord.6" AT %I3810.6 : Bool;   // Bit_06_SETPOINT
   "Carrier_69_G120DControlWord.7" AT %I3810.7 : Bool;   // Bit_07_RESET
   "Carrier_69_G120DControlWord.8" AT %I3811.0 : Bool;   // Bit_08_JOG_R
   "Carrier_69_G120DControlWord.9" AT %I3811.1 : Bool;   // Bit_09_JOG_L
   "Carrier_69_G120DControlWord.10" AT %I3811.2 : Bool;   // Bit_10_CONTR_PLC
   "Carrier_69_G120DControlWord.11" AT %I3811.3 : Bool;   // Bit_11_REVERSE
   "Carrier_69_G120DControlWord.12" AT %I3811.4 : Bool;   // Bit_12_BRAKE_RELEASE
   "Carrier_69_G120DControlWord.13" AT %I3811.5 : Bool;   // Bit_13_DDS
   "Carrier_69_G120DControlWord.14" AT %I3811.6 : Bool;   // Bit_14_DO0
   "Carrier_69_G120DControlWord.15" AT %I3811.7 : Bool;   // Bit_15_DO1
   "Carrier_69_G120DStatusWord" AT %IW3812 : Word;   // G120D_ZSW1_STATUS
   "Carrier_69_G120DStatusWord.0" AT %I3812.0 : Bool;   // Bit_00_READY_RUN
   "Carrier_69_G120DStatusWord.1" AT %I3812.1 : Bool;   // Bit_01_READY_ON
   "Carrier_69_G120DStatusWord.2" AT %I3812.2 : Bool;   // Bit_02_ENABLE
   "Carrier_69_G120DStatusWord.3" AT %I3812.3 : Bool;   // Bit_03_FAULT
   "Carrier_69_G120DStatusWord.4" AT %I3812.4 : Bool;   // Bit_04_OFF2
   "Carrier_69_G120DStatusWord.5" AT %I3812.5 : Bool;   // Bit_05_OFF3
   "Carrier_69_G120DStatusWord.6" AT %I3812.6 : Bool;   // Bit_06_LOCK_OUT
   "Carrier_69_G120DStatusWord.7" AT %I3812.7 : Bool;   // Bit_07_WARN
   "Carrier_69_G120DStatusWord.8" AT %I3813.0 : Bool;   // Bit_08_NO_DEVIATION
   "Carrier_69_G120DStatusWord.9" AT %I3813.1 : Bool;   // Bit_09_CONTR_PLC
   "Carrier_69_G120DStatusWord.10" AT %I3813.2 : Bool;   // Bit_10_F_MAX
   "Carrier_69_G120DStatusWord.11" AT %I3813.3 : Bool;   // Bit_11_LIMIT_REACHED
   "Carrier_69_G120DStatusWord.12" AT %I3813.4 : Bool;   // Bit_12_BRAKE_OPEN
   "Carrier_69_G120DStatusWord.13" AT %I3813.5 : Bool;   // Bit_13_NO_OVERTEMP
   "Carrier_69_G120DStatusWord.14" AT %I3813.6 : Bool;   // Bit_14_CW_CCW
   "Carrier_69_G120DStatusWord.15" AT %I3813.7 : Bool;   // Bit_15_OVERL
   "Carrier_69_Slot2_Input" AT %IW3814 : Word;   // SLOT 2 INPUT WORD
   "Carrier_69_CrashDetectSW" AT %I3814.0 : Bool;   // CRASH DETECT SW
   "Carrier_69_SpareSafetyInput(2_1)" AT %I3814.1 : Bool;   // SPARE SAFETY INPUT
   "Carrier_69_SpareSafetyInput(2_2)" AT %I3814.2 : Bool;   // SPARE SAFETY INPUT
   "Carrier_69_SpareSafetyInput(2_3)" AT %I3814.3 : Bool;   // SPARE SAFETY INPUT
   "Carrier_69_SpareSafetyInput(2_4)" AT %I3814.4 : Bool;   // SPARE SAFETY INPUT
   "Carrier_69_SpareSafetyInput(2_5)" AT %I3814.5 : Bool;   // SPARE SAFETY INPUT
